        [62].13   // SPARE
        [60].8   // PANEL W3 SPONGE UNIT AUTO Sw. Pos.
        [60].9   // PANEL W3 SPONGE UNIT MANUAL Sw. Pos.
        [60].10   // PANEL W3 SPONGE UNIT ON Sw. Pos.
        [60].11   // PANEL W3 SPONGE UNIT OFF Sw. Pos.
        [60].12   // PANEL W3 AIR KNIFE AUTO Sw. Pos.
        [60].13   // PANEL W3 AIR KNIFE MANUAL Sw. Pos.
        [62].9   // SPARE
        [61].0   // PANEL W3 BRUSH #1 UPPER BRUSH CONVERGE Sw. Pos.
        [61].1   // PANEL W3 BRUSH #1 UPPER BRUSH RETRACT Sw. Pos.
        [61].4   // PANEL W3 SPONGE UNIT UPPER SPONGE CONVERGE Sw. Pos.
        [61].5   // PANEL W3 SPONGE UNIT UPPER SPONGE RETRACT Sw. Pos.
        [61].6   // PANEL W3 BRUSH #1 LOWER BRUSH CONVERGE Sw. Pos.
        [61].7   // PANEL W3 BRUSH #1 LOWER BRUSH RETRACT Sw. Pos.
        [61].10   // PANEL W3 SPONGE UNIT LOWER SPONGE CONVERGE Sw. Pos.
        [61].11   // PANEL W3 SPONGE UNIT LOWER SPONGE RETRACT Sw. Pos.
        [61].12   // PANEL W3 AIR KNIFE UNIT #1 CONVERGE Sw. Pos.
        [61].13   // PANEL W3 AIR KNIFE UNIT #1 RETRACT Sw. Pos.
        [61].14   // PANEL W3 AIR KNIFE UNIT #2 CONVERGE Sw. Pos.
        [61].15   // PANEL W3 AIR KNIFE UNIT #2 RETRACT Sw. Pos.
        [62].0   // PANEL W3 Cross break Reset Push-button
        [62].1   // PANEL W3 WATER SPRAYERS AUTO Sw. Pos.
        [62].2   // PANEL W3 WATER SPRAYERS MANUAL Sw. Pos.
        [62].3   // PANEL W3 WATER SPRAYERS ON Sw. Pos.
        [62].4   // PANEL W3 WATER SPRAYERS OFF Sw. Pos.
        [64].1   // VMCC M1 DC Input Power ON
        [64].2   // VMCC M1 DC Output Power ON
        [64].4   // VMCC M1 E-STOP Power ON
        [64].5   // VMCC M1 DC Power Supply #1 ON
        [64].6   // VMCC M1 DC Power Supply #2 ON
        [64].8   // VMCC M1 Alarm Silence
        [64].9   // VMCC M1 Alarm Reset
        [64].10   // VMCC M1 E-Stop Circuit Energized
        [64].11   // VMCC M1 Crusher Bar Lowered
        [64].12   // VMCC M1 Crusher Bar Raised
        [64].13   // VMCC M1 Crusher #1 Auto mode ON=AUTO OFF=MAN
        [64].14   // VMCC M1 Crusher #1 Manual raise
        [64].15   // VMCC M1 Crusher #1 Manual lower
        [65].0   // VMCC M1 Crusher #1 Drive Fault
        [65].1   // VMCC M1 Drive Alarm Light is ON
        [65].3   // VMCC M1 Crusher #1 Test Pushbutton
        [65].4   // No. 1 Crusher Chip Blower Start Pushbutton (Top)
        [65].5   // No. 1 Crusher Chip Blower Start Pushbutton (VMCC M1)
        [65].6   // No. 1 Crusher Chip Blower Stop Pushbutton (Top)
        [65].7   // No. 1 Crusher Chip Blower Stop Pushbutton (VMCC M1)
        [65].8   // VMCC M1 SPARE
        [65].12   // VMCC M1 Crusher #1 Start Pushbutton
        [65].13   // VMCC M1 Crusher #1 Stop Pushbutton
        [65].15   // VMCC M1 Generator Running bit
        [71].2   // MB -->> Cullet M47B Run Fwd Signal
        [71].3   // MB -->> Cullet M47B Run Rev Signal
        [80].0   // NO. 1 CRUSHER Signal from Reliance drive System E-STOP
        [80].1   // NO. 1 CRUSHER Signal from C.T. master drive System DRIVE FAULT
        [80].3   // IAL TEMPERATURE ALARM
        [80].4   // Lehr Conv AUX 1 Healthy Relay
        [80].5   // Lehr Conv AUX 2 Healthy Relay
        [80].6   // Lehr Conv AUX 3 Healthy Relay
        [80].7   // Lehr Conv AUX 4 Healthy Relay
        [80].8   // Lehr Conv AUX 5 Healthy Relay
        [80].9   // Lehr Conv AUX 6 Healthy Relay
        [80].10   // Lehr Conv AUX 7 Healthy Relay
        [80].11   // Lehr Conv AUX 8 Healthy Relay
        [80].12   // Lehr Conv AUX 9 Healthy Relay
        [80].13   // Lehr Conv AUX 10 Healthy Relay
        [80].14   // Lehr Conv AUX 11 Healthy Relay
        [80].15   // Lehr Conv AUX 12 Healthy Relay
        [81]   // AUTOMAX Lehr speed Received from AutoMax
        [83].0   // Lehr Conv AUX 13 Healthy Relay
        [83].1   // Lehr Conv AUX 14 Healthy Relay
        [83].2   // Lehr Conv AUX 15 Healthy Relay
        [83].3   // Lehr Conv AUX 16 Healthy Relay
        [83].4   // Lehr Conv AUX 17 Healthy Relay
        [112].1   // Cullet -->> MB M47B Conv Fwd Signal
        [112].2   // Cullet -->> MB M47B Conv Rev Signal
        [112].3   // Cullet -->> MB M37B Conv Fwd Signal
        [112].4   // Cullet -->> MB M37B Conv Rev Signal
        [113].1   // Cullet --> MB Panel C4 Equipment Fault or Failure
        [113].2   // Cullet --> MB Panel C1 Equipment Fault or Failure
        [113].3   // Cullet --> MB Panel C2 Equipment Fault or Failure
        [113].4   // Cullet --> MB Panel C3 Equipment Fault or Failure
        [121].1   // M2 -->> MB Crusher No. 4 Is Operating
        [121].2   // M2 -->> MB Crusher No. 3 is Operating
        [121].3   // M2 ---->> MB Crusher No. 2 Is Operating
        [123].0   // M2 -->> MB Drop #1 Crusher Pushbutton
        [123].1   // M2 -->> MB Trim deck E-stop
        [123].2   // M2 -->> MB Trim deck Drive system Critical Failure
        [123].3   // M2 -->> MB Trim deck Drive fault
        [123].4   // M2 -->> MB Mainline E-stop
        [123].6   // M2 -->> MB Mainline Drive fault
        [123].11   // M2 -->> MB Drive running M2CM01
        [123].12   // M2 -->> MB Mainline Backup to
        [123].13   // M2 -->> MB Crush-all Selector sw. Status
        [123].14   // M2 -->> MB Leg 2 Is In Sleep Mode Transfer Unavailable
        [123].15   // M2 -->> MB Leg 3 Is In Sleep Mode Transfer Unavailable
        [124].0   // M2 -->> MB Leg 4 Is In Sleep Mode Transfer Unavailable
        [124].1   // M2 -->> MB Leg 5 Is In Sleep Mode Transfer Unavailable
        [124].2   // M2 -->> MB ML is in Sleep Mode
        [124].3   // M2-->Mb UL Crusher Is Faulted
        [124].4   // M2-->MB VISION SYS Rejected Plate Alarm Horn
        [127].4   // M2-->MB Float Glass Prodution
        [123]   // M2 --> MB
        [65]   // VMCC M1 Crusher
        [113]   // Cullet --> MB
        [112]   // Cullet --> MB
        [64]   // VMCC M1 INPUTS
        [121].7   // M2 -->> MB ???
        [64].0   // VMCC M1 Drive Contactor Energized
        [28].13   // CRSSBRK ZONE 3 Adapter power ON
        [30].0   // CRSSBRK ZONE 4 North Outside Bypass Switch
        [28].14   // CRSSBRK ZONE 3 Input power ON
        [124]   // M2 --> MB
        [57]   // PANEL W2
        [34].10   // MANUAL INSPCTN MODE MAN
        [34].11   // MANUAL INSPCTN MODE AUTO
        [30].9   // IMAGE AUTO Retro Reflector
        [114]   // Cullet --> MB
        [115]   // Cullet --> MB
        [80]   // LEHR Conv Healthy Relays
        [116]   // Cullet --> MB
        [117]   // Cullet --> MB
        [56]   // PANEL W2
        [125]   // M2 --> MB
        [83]   // LEHR Conv Healthy Relays
        [118]   // Cullet --> MB
        [119]   // Cullet --> MB
        [43]   // VMCC W1
        [71]   // MB --> Cullet
        [42]   // VMCC W1
        [30]   // IMAGE AUTO CRSSBRK ZONE 4
        [32]   // APC CRSSBRK ZONE 5
        [18]   // APC
        [19]   // PROCESS STOP
        [121]   // M2 --> MB
        [61]   // PANEL W3
        [60]   // PANEL W3
        [30].6   // CRSSBRK ZONE 4 South Outside Photo-cell
        [30].7   // CRSSBRK ZONE 4 South Inside Photo-cell
        [30].8   // IMAGE AUTO Open Graticule Selector Switch (UP)
        [30].14   // IMAGE AUTO Close Graticule Selector Switch (DOWN)
        [30].11   // IMAGE AUTO Cover close Acknowledge Push-button (Silence)
        [34].2   // MANUAL INSPCTN Quality defect switch (Enable/Inhibit)
        [122]   // M2 --> MB
        [28]   // CRSSBRK ZONE 3
        [30].2   // CRSSBRK ZONE 4 South Outside Bypass Switch
        [30].3   // CRSSBRK ZONE 4 South Inside Bypass Switch
        [28].15   // CRSSBRK ZONE 3 Output power ON
        [30].4   // CRSSBRK ZONE 4 North Outside Photo-cell
        [56].14   // SPARE
        [127]   // M2 --> MB
        [26]   // CRSSBRK ZONE 2
        [126]   // M2 --> MB
        [17]   // Water
        [16]   // ISRA 5D
        [3]   // PROCESS STOP
        [24]   // CRSSBRK ZONE 1
        [62]   // PANEL W3
        [26].13   // CRSSBRK ZONE 2 Adapter power ON
        [33]   // APC
        [58]   // PANEL W2
        [12]   // Bridge
        [26].15   // CRSSBRK ZONE 2 Output power ON
        [26].14   // CRSSBRK ZONE 2 Input power ON
        [30].5   // CRSSBRK ZONE 4 North Inside Photo-cell
        [30].1   // CRSSBRK ZONE 4 North Inside Bypass Switch
        [18].0   // SPARE (MARKING BRIDGE On/Off Selector switch 0=off 1=on)
        [18].1   // SPARE (MARKING BRIDGE Auto/Manual 0=Manual 1=Auto)
        [16].2   // Spare
        [16].11   // Spare
        [16].12   // Spare
        [16].13   // Spare
        [16].15   // Spare
        [17].0   // Spare
        [17].6   // Spare
        [17].8   // Spare
        [17].12   // SPARE (Chilled Water Blower VFD Is At Speed)
        [17].15   // SPARE (ROCKWELL CAPPING SYSTEM: 50mm of Glass Travel Pulse Signal)
        [33].9   // SPARE (Apc system 0ff)
        [34]   // LOW-E MAUAL INSPCTN (MI_6CS)
        [43].4   // VMCC W1 Upper Sponge Drive fault (NOT USED ANYMORE)
        [43].5   // VMCC W1 Lower Sponge Drive fault (NOT USED ANYMORE)
        [42].1   // VMCC W1 Drive Contactor Energized (NOT USED ANYMORE)
        [42].2   // VMCC W1 DC Input Power ON (NOT USED ANYMORE)
        [42].3   // VMCC W1 DC Output Power ON (NOT USED ANYMORE)
        [42].5   // VMCC W1 E-STOP Power ON (NOT USED ANYMORE)
        [42].6   // VMCC W1 DC Power Supply #1 ON (NOT USED ANYMORE)
        [42].7   // VMCC W1 DC Power Supply #2 ON (NOT USED ANYMORE)
        [42].8   // VMCC W1 Alarm Silence (NOT USED ANYMORE)
        [42].10   // VMCC W1 E-STOP ACTIVE (NOT USED ANYMORE)
        [42].11   // VMCC W1 Drive Comm. Power (NOT USED ANYMORE)
        [43].12   // VMCC W1 Crusher #1 Start Pushbutton (NOT USED ANYMORE)
        [43].13   // VMCC W1 Crusher #1 Stop Pushbutton (NOT USED ANYMORE)
        [56].4   // PANEL W2 BRUSH #2 AUTO Sw. Pos. (NOT USED ANYMORE)
        [56].5   // PANEL W2 BRUSH #2 MANUAL Sw. Pos. (NOT USED ANYMORE)
        [56].6   // PANEL W2 BRUSH #2 ON Sw. Pos. (NOT USED ANYMORE)
        [56].7   // PANEL W2 BRUSH #2 OFF Sw. Pos. (NOT USED ANYMORE)
        [57].2   // PANEL W2 BRUSH #2 UPPER BRUSH CONVERGE Sw. Pos. (NOT USED ANYMORE)
        [57].3   // PANEL W2 BRUSH #2 UPPER BRUSH RETRACT Sw. Pos. (NOT USED ANYMORE)
        [57].8   // PANEL W2 BRUSH #2 LOWER BRUSH CONVERGE Sw. Pos. (NOT USED ANYMORE)
        [57].9   // PANEL W2 BRUSH #2 LOWER BRUSH RETRACT Sw. Pos. (NOT USED ANYMORE)
        [60].4   // PANEL W3 BRUSH #2 AUTO Sw. Pos. (NOT USED ANYMORE)
        [60].5   // PANEL W3 BRUSH #2 MANUAL Sw. Pos. (NOT USED ANYMORE)
        [60].6   // PANEL W3 BRUSH #2 ON Sw. Pos. (NOT USED ANYMORE)
        [60].7   // PANEL W3 BRUSH #2 OFF Sw. Pos. (NOT USED ANYMORE)
        [61].2   // PANEL W3 BRUSH #2 UPPER BRUSH CONVERGE Sw. Pos. (NOT USED ANYMORE)
        [61].3   // PANEL W3 BRUSH #2 UPPER BRUSH RETRACT Sw. Pos. (NOT USED ANYMORE)
        [61].8   // PANEL W3 BRUSH #2 LOWER BRUSH CONVERGE Sw. Pos. (NOT USED ANYMORE)
        [61].9   // PANEL W3 BRUSH #2 LOWER BRUSH RETRACT Sw. Pos. (NOT USED ANYMORE)
        [58].5   // PANEL W2 SELECTOR SWITCH CITRIC ACID WASHER ON (# W2) (NOT USED ANYMORE)
        [58].6   // PANEL W2 SELECTOR SWITCH CITRIC ACID WASHER OFF (# W2) (NOT USED ANYMORE)
        [62].5   // PANEL W3 SELECTOR SWITCH CITRIC ACID WASHER ON (# W3) (NOT USED ANYMORE)
        [62].6   // PANEL W3 SELECTOR SWITCH CITRIC ACID WASHER OFF (# W3) (NOT USED ANYMORE)
        [113].0   // Cullet --> MB SYSTEM LOCAL HEARTBEAT FOR HOST PLC
        [113].5   // Cullet --> MB FIX MMI M-47B Conveyor Running Reverse
        [114].1   // LEG 4 EOL FEEDER AUTO RUN STATUS
        [114].2   // LEG 5 EOL FEEDER AUTO RUN STATUS
        [114].3   // PANEL C4 - TRIM DROP VP 917078 Running at Speed
        [114].4   // PANEL C3 - CR#3 VP 917067 VFD FAULT STATUS
        [114].5   // PANEL C3 - CR#3 VP 917067 VFD RUNNING STATUS
        [114].6   // PANEL C3 M34T TO M34 TRANS VP 917066 VFD FAULT STATUS
        [114].7   // PANEL C3 M34T TO M34 TRANS VP 917066 VFD RUNNING STATUS
        [114].10   // PANEL C3 VP 917070 VFD FAULT STATUS
        [114].11   // PANEL C3 VP 917070 VFD RUNNING STATUS
        [114].12   // PANEL C3 VP 917071 VFD FAULT STATUS
        [114].13   // PANEL C3 VP 917071 VFD RUNNING STATUS
        [114].14   // PANEL C2 VP 917077 VFD FAULT STATUS
        [114].15   // PANEL C2 VP 917077 VFD RUNNING STATUS
        [115].0   // PANEL C4 M34T MAIN #1 CONV RUNNING STATUS
        [115].1   // LEG 3 EOL FEEDER AUTO RUN STATUS
        [115].2   // PANEL C4 M-32 CONVEYOR RUNNING STATUS
        [115].3   // PANEL C4 M-33 CONVEYOR RUNNING STATUS
        [115].4   // PANEL C4 M34T MAIN #1 CONV E-STOP STATUS
        [115].6   // PANEL C4 M-32 CONVEYOR E-STOP STATUS
        [115].7   // PANEL C4 M-33 CONVEYOR E-STOP STATUS
        [115].8   // PANEL C4 M34T MAIN CONV #1 ZERO SPEED STATUS
        [115].10   // PANEL C4 M-32 CONVEYOR ZERO SPEED SWITCH STATUS
        [115].11   // PANEL C4 M-33 CONVEYOR ZERO SPEED STATUS
        [115].12   // PANEL C2 VP 917076 VFD FAULT STATUS
        [115].13   // PANEL C2 VP 917076 VFD RUNNING STATUS
        [115].14   // PANEL C2 VP 917075 VFD FAULT STATUS
        [115].15   // PANEL C2 VP 917075 VFD RUNNING STATUS
        [116].0   // PANEL C4 - CR#4 VP 917068 VFD RUNNING STATUS
        [116].1   // LEG 5 FEEDER DRIVE RUNNING STATUS
        [116].2   // PANEL C2 VP 917074 VFD FAULT STATUS
        [116].3   // PANEL C2 VP 917074 VFD RUNNING STATUS
        [116].4   // PANEL C4 - CR#4 VP 917068 VFD FAULT STATUS
        [116].7   // PANEL C2 VP 917073 VFD FAULT STATUS
        [116].8   // PANEL C2 VP 917073 VFD RUNNING STATUS
        [116].9   // PANEL C2 VP 917072 VFD FAULT STATUS
        [116].10   // PANEL C2 VP 917072 VFD RUNNING STATUS
        [116].11   // PANEL C1 VP 917060 VFD FAULT STATUS
        [116].12   // PANEL C1 VP 917060 VFD RUNNING STATUS
        [116].13   // PANEL C3 M-40 CONVEYOR RUNNING STATUS
        [116].14   // PANEL C3 M-40 CONVEYOR E-STOP STATUS
        [116].15   // PANEL C3 M-40 CONVEYOR ZERO SPEED SWITCH STATUS
        [117].0   // M47A_RUN_STAT PANEL C1 M-47A CONVEYOR RUNNING STATUS
        [117].1   // M47A_ESTOP_STAT PANEL C1 M-47A CONVEYOR E-STOP STATUS
        [117].2   // M47A_ZSS_STAT PANEL C1 M-47A CONVEYOR ZERO SPEED SWITCH STATUS
        [117].3   // M47B_RUN_STAT PANEL C1 M-47B CONVEYOR RUNNING STATUS
        [117].4   // M47B_ESTOP_STAT PANEL C1 M-47B CONVEYOR E-STOP STATUS
        [117].5   // M47B_ZSS_STAT PANEL C1 M-47B CONVEYOR ZERO SPEED SWITCH STATUS
        [117].6   // M46_RUN_STAT PANEL C1 M-46 CONVEYOR RUNNING STATUS
        [117].7   // M46_ESTOP_STAT PANEL C1 M-46 CONVEYOR E-STOP STATUS
        [117].8   // M46_ZSS_STAT PANEL C1 M-46 CONVEYOR ZERO SPEED SWITCH STATUS
        [117].9   // M45B_RUN_STAT PANEL C1 M-45B CONVEYOR RUNNING STATUS
        [117].10   // M45B_ESTOP_STAT PANEL C1 M-45B CONVEYOR E-STOP STATUS
        [117].11   // M45B_ZSS_STAT PANEL C1 M-45B CONVEYOR ZERO SPEED SWITCH STATUS
        [117].12   // M37A_RUN_STAT PANEL C2 M-37A CONVEYOR RUNNING STATUS
        [117].13   // M37A_ESTOP_STAT PANEL C2 M-37A CONVEYOR E-STOP STATUS
        [117].14   // M37A_ZSS_STAT PANEL C2 M-37A CONVEYOR ZERO SPEED SWITCH STATUS
        [117].15   // M37B_RUN_STAT PANEL C2 M-37B CONVEYOR RUNNING STATUS
        [118].0   // M37B_ESTOP_STAT PANEL C2 M-37B CONVEYOR E-STOP STATUS
        [118].1   // M37B_ZSS_STAT PANEL C2 M-37B CONVEYOR ZERO SPEED SWITCH STATUS
        [118].2   // M36_RUN_STAT PANEL C2 M-36 CONVEYOR RUNNING STATUS
        [118].3   // M36_ESTOP_STAT PANEL C2 M-36 CONVEYOR E-STOP STATUS
        [118].4   // M36_ZSS_STAT PANEL C2 M-36 CONVEYOR ZERO SPEED SWITCH STATUS
        [118].5   // M35_RUN_STAT PANEL C2 M-35 CONVEYOR RUNNING STATUS
        [118].6   // M35_ESTOP_STAT PANEL C2 M-35 CONVEYOR E-STOP STATUS
        [118].7   // M35_ZSS_STAT PANEL C2 M-35 CONVEYOR ZERO SPEED SWITCH STATUS
        [118].8   // CHPR_RUN_STAT PANEL C2 CHOPPER 917014 RUNNING STATUS
        [118].9   // CHPR_ESTOP_STAT PANEL C2 CHOPPER 917014 E-STOP STATUS
        [118].10   // CHPR_ZSS_STAT PANEL C2 CHOPPER 917014 ZERO SPEED SWITCH STATUS
        [118].11   // M45_RUN_STAT PANEL C2 M-45 CONVEYOR RUNNING STATUS
        [118].12   // M45_ESTOP_STAT PANEL C2 M-45 CONVEYOR E-STOP STATUS
        [118].13   // M45_ZSS_STAT PANEL C2 M-45 CONVEYOR ZERO SPEED SWITCH STATUS
        [118].14   // M45A_RUN_STAT PANEL C2 M-45A CONVEYOR RUNNING STATUS
        [118].15   // M45A_ESTOP_STAT PANEL C2 M-45A CONVEYOR E-STOP STATUS
        [119].0   // M45A_ZSS_STAT PANEL C2 M-45A CONVEYOR ZERO SPEED SWITCH STATUS
        [119].1   // M34_RUN_STAT PANEL C3 M-34 CONVEYOR RUNNING STATUS
        [119].2   // M34_ESTOP_STAT PANEL C3 M-34 CONVEYOR E-STOP STATUS
        [119].3   // M34_ZSS_STAT PANEL C3 M-34 CONVEYOR ZERO SPEED SWITCH STATUS
        [119].4   // M44_RUN_STAT PANEL C3 M-44 CONVEYOR RUNNING STATUS
        [119].5   // M44_ESTOP_STAT PANEL C3 M-44 CONVEYOR E-STOP STATUS
        [119].6   // M44_ZSS_STAT PANEL C3 M-44 CONVEYOR ZERO SPEED SWITCH STATUS
        [119].7   // M43_RUN_STAT PANEL C3 M-43 CONVEYOR RUNNING STATUS
        [119].8   // M43_ESTOP_STAT PANEL C3 M-43 CONVEYOR E-STOP STATUS
        [119].9   // M43_ZSS_STAT PANEL C3 M-43 CONVEYOR ZERO SPEED SWITCH STATUS
        [119].10   // M41_RUN_STAT PANEL C3 M-41 CONVEYOR RUNNING STATUS
        [119].11   // M41_ESTOP_STAT PANEL C3 M-41 CONVEYOR E-STOP STATUS
        [119].12   // M41_ZSS_STAT PANEL C3 M-41 CONVEYOR ZERO SPEED SWITCH STATUS
        [119].13   // M42_RUN_STAT PANEL C3 M-42 CONVEYOR RUNNING STATUS
        [119].14   // M42_ESTOP_STAT PANEL C3 M-42 CONVEYOR E-STOP STATUS
        [119].15   // M42_ZSS_STAT PANEL C3 M-42 CONVEYOR ZERO SPEED SWITCH STATUS
   IA_ACK_PB : ALIAS FOR I[30].11;
   IA_CLOSE_GRAT : ALIAS FOR I[30].14;
   IA_COVER_CLOSED : ALIAS FOR N54[281].5;
   IA_COVER_VLVE : ALIAS FOR O[31].10;
   IA_GRAT_OPEN_SS : ALIAS FOR I[30].8;
   IA_RET_CL_PROX : ALIAS FOR I[30].12;
   IA_RET_CLSD_ACK : ALIAS FOR N54[281].6;
   INDEX : ALIAS FOR S[24];
   INIT_TIMER : ALIAS FOR T4[0];
   IW_FE1_BTR : ALIAS FOR W_N7[32];
   LEG2_SLEEP : ALIAS FOR I[123].14;
   LEG3_SLEEP : ALIAS FOR I[123].15;
   LEG4_SLEEP : ALIAS FOR I[124].0;
   LEG5_SLEEP : ALIAS FOR I[124].1;
   LEHR_2IN_PULSE : ALIAS FOR B73[0].1;
   LEHR_SPEED : ALIAS FOR N60[1];
   LEHRSPD_AUTOMAX : ALIAS FOR N98[1];
   LEHRSPD_AVE : ALIAS FOR N98[2];
   LEHRSPD_CURRENT : ALIAS FOR N98[5];
   LEHRSPD_STD : ALIAS FOR N98[3];
   M1_ALM_FLT_RLY : ALIAS FOR O[66].13;
   M1_ALM_RESET : ALIAS FOR I[64].9;
   M1_ALM_SILENCE : ALIAS FOR I[64].8;
   M1_DC_INPOW : ALIAS FOR I[64].1;
   M1_DC_OUTPOW : ALIAS FOR I[64].2;
   M1_DC_PS1 : ALIAS FOR I[64].5;
   M1_DC_PS2 : ALIAS FOR I[64].6;
   M1_DRV_CONT_ON : ALIAS FOR I[64].0;
   M1_ESTOP_ON : ALIAS FOR I[64].10;
   M1_ESTOPPOW : ALIAS FOR I[64].4;
   M202_M1_DR : AXIS_CIP_DRIVE; {access Read Only}
   M202_M1_DR_IN_MAJ : MOTION_INSTRUCTION := (FLAGS := 570425344, DN := 1); {access None}
   M202_M1_DR_IN_MAM : MOTION_INSTRUCTION := (FLAGS := 33554432); {access None}
   M202_M1_DR_IN_MAR : MOTION_INSTRUCTION := (FLAGS := 33554432); {access None}
   M202_M1_DR_IN_MAS : MOTION_INSTRUCTION := (FLAGS := -1442840576, EN := 1, DN := 1, PC := 1); {access None}
   M202_M1_DR_IN_MCD : MOTION_INSTRUCTION := (FLAGS := 570425344, DN := 1); {access None}
   M202_M1_DR_IN_MRP : MOTION_INSTRUCTION := (FLAGS := 33554432); {access None}
   M202_M1_DR_MAFR : MOTION_INSTRUCTION := (FLAGS := 301989888, ER := 1, ERR := 11); {access None}
   M202_M1_DR_MDR : MOTION_INSTRUCTION := (FLAGS := -1845493760, EN := 1, ER := 1, ERR := 11); {access None}
   M202_M1_DR_MSF : MOTION_INSTRUCTION := (FLAGS := 570425344, DN := 1, STATUS := 2, STATE := 1); {access None}
   M202_M1_DR_MSO : MOTION_INSTRUCTION := (FLAGS := -1610612736, EN := 1, DN := 1, STATE := 1); {access None}
   M202_M1_DR_OUT_MAJ : MOTION_INSTRUCTION := (FLAGS := 570425344, DN := 1); {access None}
   M202_M1_DR_OUT_MAM : MOTION_INSTRUCTION := (FLAGS := 33554432); {access None}
   M202_M1_DR_OUT_MAR : MOTION_INSTRUCTION := (FLAGS := 33554432); {access None}
   M202_M1_DR_OUT_MAS : MOTION_INSTRUCTION := (FLAGS := -1442840576, EN := 1, DN := 1, PC := 1); {access None}
   M202_M1_DR_OUT_MCD : MOTION_INSTRUCTION := (FLAGS := 570425344, DN := 1); {access None}
   M202_M1_DR_OUT_MRP : MOTION_INSTRUCTION := (FLAGS := 33554432); {access None}
   M203_M1_DR : AXIS_CIP_DRIVE; {access Read Only}
   M203_M1_DR_IN_MAJ : MOTION_INSTRUCTION := (FLAGS := 570425344, DN := 1); {access None}
   M203_M1_DR_IN_MAM : MOTION_INSTRUCTION := (FLAGS := 33554432); {access None}
   M203_M1_DR_IN_MAR : MOTION_INSTRUCTION := (FLAGS := 33554432); {access None}
   M203_M1_DR_IN_MAS : MOTION_INSTRUCTION := (FLAGS := -1442840576, EN := 1, DN := 1, PC := 1); {access None}
   M203_M1_DR_IN_MCD : MOTION_INSTRUCTION := (FLAGS := 570425344, DN := 1); {access None}
   M203_M1_DR_IN_MRP : MOTION_INSTRUCTION := (FLAGS := 33554432); {access None}
   M203_M1_DR_MAFR : MOTION_INSTRUCTION := (FLAGS := 301989888, ER := 1, ERR := 11); {access None}
   M203_M1_DR_MDR : MOTION_INSTRUCTION := (FLAGS := -1845493760, EN := 1, ER := 1, ERR := 11); {access None}
   M203_M1_DR_MSF : MOTION_INSTRUCTION := (FLAGS := 570425344, DN := 1, STATUS := 2, STATE := 1); {access None}
   M203_M1_DR_MSO : MOTION_INSTRUCTION := (FLAGS := -1610612736, EN := 1, DN := 1, STATE := 1); {access None}
   M203_M1_DR_OUT_MAJ : MOTION_INSTRUCTION := (FLAGS := 570425344, DN := 1); {access None}
   M203_M1_DR_OUT_MAM : MOTION_INSTRUCTION := (FLAGS := 33554432); {access None}
   M203_M1_DR_OUT_MAR : MOTION_INSTRUCTION := (FLAGS := 33554432); {access None}
   M203_M1_DR_OUT_MAS : MOTION_INSTRUCTION := (FLAGS := -1442840576, EN := 1, DN := 1, PC := 1); {access None}
   M203_M1_DR_OUT_MCD : MOTION_INSTRUCTION := (FLAGS := 570425344, DN := 1); {access None}
   M203_M1_DR_OUT_MRP : MOTION_INSTRUCTION := (FLAGS := 33554432); {access None}
   M203DROP : MAC_DROPCONV := (OUTPUT_xHLUpDownPushbutton := 1, INPUT_xProtection := 1, INPUT_xProtectionBrake := 1, AUX_tmOFFEachCutAcceleration.PRE := 2000, AUX_tmOFFEachCutAcceleration.ACC := 2000, AUX_tmOFFAcceleration.PRE := 8805, AUX_tmOFFAcceleration.ACC := 8805, AUX_tmONFeedbackMovAlarm.PRE := 2000, AUX_tmONFeedbackAlarm.PRE := 2000, AUX_tmONFeedbackBrakeAlarm.PRE := 7000, AUX_tmONMismatchSensorAlarm.PRE := 7000, AUX_tmONUpSensorAlarm.PRE := 5000, AUX_tmONDownSensorAlarm.PRE := 5000, AUX_tmONForceUp.PRE := 2000, AUX_tmONEmCutTimeout.PRE := 120000, AUX_dDistanceToDescent_cmm := 25000, AUX_dDistanceToCheckGlass_cmm := 100000, AUX_dConveyorLength_cmm := 440000, AUX_dAccelerationTime_ms := 2147483647, AUX_dAccelerationFactor := 3, AUX_dMaxSpeed_mm_min := 30000, ST_xConveyorDwRequest := 1, OSR_xCutForQltPopupEnd := 1); {access None}
   M203DROP_ALM : MAC_DROPCONV_ALM; {access Read Only}
        .rgxStoppingFaults[0].0   // Protection lifting
        .rgxStoppingFaults[0].1   // Protection brake
        .rgxStoppingFaults[0].2   // Feedback lifting
        .rgxStoppingFaults[0].3   // Feedback brake
        .rgxStoppingFaults[0].5   // A206SQ2.Timeout frame low
        .rgxStoppingFaults[0].6   // A206SQ1/2.Sensor high/low mismatch (same status)
        .rgxStoppingFaults[0].4   // A206SQ1.Timeout frame high
        .rgxStoppingFaults[0].7   // A206SQ3/4.Tilting safety bar disinsered
   M203DROP_HMR : MAC_DROPCONV_HMR := (dMode := 1, dStatus := 1, dDistanceFromSnaproll_cmm := 4190000); {access Read Only}
   M203DROP_HMW : MAC_DROPCONV_HMW := (dDistanceFromSnaproll_cmm := 4632000);
   M204_M1_DR : AXIS_CIP_DRIVE; {access Read Only}
   M204_M1_DR_IN_MAJ : MOTION_INSTRUCTION := (FLAGS := 570425344, DN := 1); {access None}
   M204_M1_DR_IN_MAM : MOTION_INSTRUCTION := (FLAGS := 33554432); {access None}
   M204_M1_DR_IN_MAR : MOTION_INSTRUCTION := (FLAGS := 33554432); {access None}
   M204_M1_DR_IN_MAS : MOTION_INSTRUCTION := (FLAGS := -1442840576, EN := 1, DN := 1, PC := 1); {access None}
   M204_M1_DR_IN_MCD : MOTION_INSTRUCTION := (FLAGS := 570425344, DN := 1); {access None}
   M204_M1_DR_IN_MRP : MOTION_INSTRUCTION := (FLAGS := 33554432); {access None}
   M204_M1_DR_MAFR : MOTION_INSTRUCTION := (FLAGS := 301989888, ER := 1, ERR := 11); {access None}
   M204_M1_DR_MDR : MOTION_INSTRUCTION := (FLAGS := -1845493760, EN := 1, ER := 1, ERR := 11); {access None}
   M204_M1_DR_MSF : MOTION_INSTRUCTION := (FLAGS := 570425344, DN := 1, STATUS := 2, STATE := 1); {access None}
   M204_M1_DR_MSO : MOTION_INSTRUCTION := (FLAGS := -1610612736, EN := 1, DN := 1, STATE := 1); {access None}
   M204_M1_DR_OUT_MAJ : MOTION_INSTRUCTION := (FLAGS := 570425344, DN := 1); {access None}
   M204_M1_DR_OUT_MAM : MOTION_INSTRUCTION := (FLAGS := 33554432); {access None}
   M204_M1_DR_OUT_MAR : MOTION_INSTRUCTION := (FLAGS := 33554432); {access None}
   M204_M1_DR_OUT_MAS : MOTION_INSTRUCTION := (FLAGS := -1442840576, EN := 1, DN := 1, PC := 1); {access None}
   M204_M1_DR_OUT_MCD : MOTION_INSTRUCTION := (FLAGS := 570425344, DN := 1); {access None}
   M204_M1_DR_OUT_MRP : MOTION_INSTRUCTION := (FLAGS := 33554432); {access None}
   M205BREAKER : MAC_BREAKER := (ST_xBreakerRunningRequest := 1, OSR_xBreakerRunning := 1, INPUT_xProtectionFan := 1, INPUT_xStopBreaker := 1, INPUT_xThermalProbe := 1, OUTPUT_xBreakerRun := 1, AUX_tmONCrusherStopDelayed.PRE := 320000, AUX_tmONFeedbackBreakerRot.PRE := 15000, AUX_tmONBreakControlRotation.PRE := 5000, AUX_tmONFeedbackBrakeBreakRot.PRE := 2000, AUX_tmONFeedbackExclusionInduct.PRE := 5000); {access None}
   M205BREAKER_ALM : MAC_BREAKER_ALM; {access Read Only}
        .rgxStoppingFaults[0].5   // Exclusion inductance feedback
        .rgxStoppingFaults[0].3   // Drive error
        .rgdCodeAlarm[0]   // A60AZ1.Error Code
        .rgxStoppingFaults[0].2   // Motor thermal probe
        .rgxStoppingFaults[0].4   // A56QS1.Safety motor sectioning
        .rgxStoppingFaults[0].0   // Rotation feedback
        .rgxStoppingFaults[0].1   // Protection rotation
        .rgxStoppingFaults[0].6   // A207SQ1.Breaker rotation sensor
        .rgxFaults[0].0   // A63QM2.Protection fan rotation
   M205BREAKER_HMR : MAC_BREAKER_HMR := (dBreakerStatus := 1); {access Read Only}
   M205BREAKER_HMW : MAC_BREAKER_HMW := (dTimeoutRunningCrusher_ms := 320000);
   M206_M1_DR : AXIS_CIP_DRIVE; {access Read Only}
   M206_M1_DR_IN_MAJ : MOTION_INSTRUCTION := (FLAGS := 570425344, DN := 1); {access None}
   M206_M1_DR_IN_MAM : MOTION_INSTRUCTION := (FLAGS := 33554432); {access None}
   M206_M1_DR_IN_MAR : MOTION_INSTRUCTION := (FLAGS := 33554432); {access None}
   M206_M1_DR_IN_MAS : MOTION_INSTRUCTION := (FLAGS := -1442840576, EN := 1, DN := 1, PC := 1); {access None}
   M206_M1_DR_IN_MCD : MOTION_INSTRUCTION := (FLAGS := 570425344, DN := 1); {access None}
   M206_M1_DR_IN_MRP : MOTION_INSTRUCTION := (FLAGS := 33554432); {access None}
   M206_M1_DR_MAFR : MOTION_INSTRUCTION := (FLAGS := 301989888, ER := 1, ERR := 11); {access None}
   M206_M1_DR_MDR : MOTION_INSTRUCTION := (FLAGS := -1845493760, EN := 1, ER := 1, ERR := 11); {access None}
   M206_M1_DR_MSF : MOTION_INSTRUCTION := (FLAGS := 570425344, DN := 1, STATUS := 2, STATE := 1); {access None}
   M206_M1_DR_MSO : MOTION_INSTRUCTION := (FLAGS := -1610612736, EN := 1, DN := 1, STATE := 1); {access None}
   M206_M1_DR_OUT_MAJ : MOTION_INSTRUCTION := (FLAGS := 570425344, DN := 1); {access None}
   M206_M1_DR_OUT_MAM : MOTION_INSTRUCTION := (FLAGS := 33554432); {access None}
   M206_M1_DR_OUT_MAR : MOTION_INSTRUCTION := (FLAGS := 33554432); {access None}
   M206_M1_DR_OUT_MAS : MOTION_INSTRUCTION := (FLAGS := -1442840576, EN := 1, DN := 1, PC := 1); {access None}
   M206_M1_DR_OUT_MCD : MOTION_INSTRUCTION := (FLAGS := 570425344, DN := 1); {access None}
   M206_M1_DR_OUT_MRP : MOTION_INSTRUCTION := (FLAGS := 33554432); {access None}
   M207_M1_DR : AXIS_CIP_DRIVE; {access Read Only}
   M207_M1_DR_IN_MAJ : MOTION_INSTRUCTION := (FLAGS := 570425344, DN := 1); {access None}
   M207_M1_DR_IN_MAM : MOTION_INSTRUCTION := (FLAGS := 33554432); {access None}
   M207_M1_DR_IN_MAR : MOTION_INSTRUCTION := (FLAGS := 33554432); {access None}
   M207_M1_DR_IN_MAS : MOTION_INSTRUCTION := (FLAGS := -1442840576, EN := 1, DN := 1, PC := 1); {access None}
   M207_M1_DR_IN_MCD : MOTION_INSTRUCTION := (FLAGS := 570425344, DN := 1); {access None}
   M207_M1_DR_IN_MRP : MOTION_INSTRUCTION := (FLAGS := 33554432); {access None}
   M207_M1_DR_MAFR : MOTION_INSTRUCTION := (FLAGS := 301989888, ER := 1, ERR := 11); {access None}
   M207_M1_DR_MDR : MOTION_INSTRUCTION := (FLAGS := -1845493760, EN := 1, ER := 1, ERR := 11); {access None}
   M207_M1_DR_MSF : MOTION_INSTRUCTION := (FLAGS := 570425344, DN := 1, STATUS := 2, STATE := 1); {access None}
   M207_M1_DR_MSO : MOTION_INSTRUCTION := (FLAGS := -1610612736, EN := 1, DN := 1, STATE := 1); {access None}
   M207_M1_DR_OUT_MAJ : MOTION_INSTRUCTION := (FLAGS := 570425344, DN := 1); {access None}
   M207_M1_DR_OUT_MAM : MOTION_INSTRUCTION := (FLAGS := 33554432); {access None}
   M207_M1_DR_OUT_MAR : MOTION_INSTRUCTION := (FLAGS := 33554432); {access None}
   M207_M1_DR_OUT_MAS : MOTION_INSTRUCTION := (FLAGS := -1442840576, EN := 1, DN := 1, PC := 1); {access None}
   M207_M1_DR_OUT_MCD : MOTION_INSTRUCTION := (FLAGS := 570425344, DN := 1); {access None}
   M207_M1_DR_OUT_MRP : MOTION_INSTRUCTION := (FLAGS := 33554432); {access None}
   M208_M1_DR : AXIS_CIP_DRIVE; {access Read Only}
   M208_M1_DR_IN_MAJ : MOTION_INSTRUCTION := (FLAGS := 570425344, DN := 1); {access None}
   M208_M1_DR_IN_MAM : MOTION_INSTRUCTION := (FLAGS := 33554432); {access None}
   M208_M1_DR_IN_MAR : MOTION_INSTRUCTION := (FLAGS := 33554432); {access None}
   M208_M1_DR_IN_MAS : MOTION_INSTRUCTION := (FLAGS := -1442840576, EN := 1, DN := 1, PC := 1); {access None}
   M208_M1_DR_IN_MCD : MOTION_INSTRUCTION := (FLAGS := 570425344, DN := 1); {access None}
   M208_M1_DR_IN_MRP : MOTION_INSTRUCTION := (FLAGS := 33554432); {access None}
   M208_M1_DR_MAFR : MOTION_INSTRUCTION := (FLAGS := 301989888, ER := 1, ERR := 11); {access None}
   M208_M1_DR_MDR : MOTION_INSTRUCTION := (FLAGS := -1845493760, EN := 1, ER := 1, ERR := 11); {access None}
   M208_M1_DR_MSF : MOTION_INSTRUCTION := (FLAGS := 570425344, DN := 1, STATUS := 2, STATE := 1); {access None}
   M208_M1_DR_MSO : MOTION_INSTRUCTION := (FLAGS := -1610612736, EN := 1, DN := 1, STATE := 1); {access None}
   M208_M1_DR_OUT_MAJ : MOTION_INSTRUCTION := (FLAGS := 570425344, DN := 1); {access None}
   M208_M1_DR_OUT_MAM : MOTION_INSTRUCTION := (FLAGS := 33554432); {access None}
   M208_M1_DR_OUT_MAR : MOTION_INSTRUCTION := (FLAGS := 33554432); {access None}
   M208_M1_DR_OUT_MAS : MOTION_INSTRUCTION := (FLAGS := -1442840576, EN := 1, DN := 1, PC := 1); {access None}
   M208_M1_DR_OUT_MCD : MOTION_INSTRUCTION := (FLAGS := 570425344, DN := 1); {access None}
   M208_M1_DR_OUT_MRP : MOTION_INSTRUCTION := (FLAGS := 33554432); {access None}
   M209_M1_DR : AXIS_CIP_DRIVE; {access Read Only}
   M209_M1_DR_IN_MAJ : MOTION_INSTRUCTION := (FLAGS := 570425344, DN := 1); {access None}
   M209_M1_DR_IN_MAM : MOTION_INSTRUCTION := (FLAGS := 33554432); {access None}
   M209_M1_DR_IN_MAR : MOTION_INSTRUCTION := (FLAGS := 33554432); {access None}
   M209_M1_DR_IN_MAS : MOTION_INSTRUCTION := (FLAGS := -1442840576, EN := 1, DN := 1, PC := 1); {access None}
   M209_M1_DR_IN_MCD : MOTION_INSTRUCTION := (FLAGS := 570425344, DN := 1); {access None}
   M209_M1_DR_IN_MRP : MOTION_INSTRUCTION := (FLAGS := 33554432); {access None}
   M209_M1_DR_MAFR : MOTION_INSTRUCTION := (FLAGS := 301989888, ER := 1, ERR := 11); {access None}
   M209_M1_DR_MDR : MOTION_INSTRUCTION := (FLAGS := -1845493760, EN := 1, ER := 1, ERR := 11); {access None}
   M209_M1_DR_MSF : MOTION_INSTRUCTION := (FLAGS := 570425344, DN := 1, STATUS := 2, STATE := 1); {access None}
   M209_M1_DR_MSO : MOTION_INSTRUCTION := (FLAGS := -1610612736, EN := 1, DN := 1, STATE := 1); {access None}
   M209_M1_DR_OUT_MAJ : MOTION_INSTRUCTION := (FLAGS := 570425344, DN := 1); {access None}
   M209_M1_DR_OUT_MAM : MOTION_INSTRUCTION := (FLAGS := 33554432); {access None}
   M209_M1_DR_OUT_MAR : MOTION_INSTRUCTION := (FLAGS := 33554432); {access None}
   M209_M1_DR_OUT_MAS : MOTION_INSTRUCTION := (FLAGS := -1442840576, EN := 1, DN := 1, PC := 1); {access None}
   M209_M1_DR_OUT_MCD : MOTION_INSTRUCTION := (FLAGS := 570425344, DN := 1); {access None}
   M209_M1_DR_OUT_MRP : MOTION_INSTRUCTION := (FLAGS := 33554432); {access None}
   M210_M1_DR : AXIS_CIP_DRIVE; {access Read Only}
   M210_M1_DR_IN_MAJ : MOTION_INSTRUCTION := (FLAGS := 570425344, DN := 1); {access None}
   M210_M1_DR_IN_MAM : MOTION_INSTRUCTION := (FLAGS := 33554432); {access None}
   M210_M1_DR_IN_MAR : MOTION_INSTRUCTION := (FLAGS := 33554432); {access None}
   M210_M1_DR_IN_MAS : MOTION_INSTRUCTION := (FLAGS := -1442840576, EN := 1, DN := 1, PC := 1); {access None}
   M210_M1_DR_IN_MCD : MOTION_INSTRUCTION := (FLAGS := 570425344, DN := 1); {access None}
   M210_M1_DR_IN_MRP : MOTION_INSTRUCTION := (FLAGS := 33554432); {access None}
   M210_M1_DR_MAFR : MOTION_INSTRUCTION := (FLAGS := 301989888, ER := 1, ERR := 11); {access None}
   M210_M1_DR_MDR : MOTION_INSTRUCTION := (FLAGS := -1845493760, EN := 1, ER := 1, ERR := 11); {access None}
   M210_M1_DR_MSF : MOTION_INSTRUCTION := (FLAGS := 570425344, DN := 1, STATUS := 2, STATE := 1); {access None}
   M210_M1_DR_MSO : MOTION_INSTRUCTION := (FLAGS := -1610612736, EN := 1, DN := 1, STATE := 1); {access None}
   M210_M1_DR_OUT_MAJ : MOTION_INSTRUCTION := (FLAGS := 570425344, DN := 1); {access None}
   M210_M1_DR_OUT_MAM : MOTION_INSTRUCTION := (FLAGS := 33554432); {access None}
   M210_M1_DR_OUT_MAR : MOTION_INSTRUCTION := (FLAGS := 33554432); {access None}
   M210_M1_DR_OUT_MAS : MOTION_INSTRUCTION := (FLAGS := -1442840576, EN := 1, DN := 1, PC := 1); {access None}
   M210_M1_DR_OUT_MCD : MOTION_INSTRUCTION := (FLAGS := 570425344, DN := 1); {access None}
   M210_M1_DR_OUT_MRP : MOTION_INSTRUCTION := (FLAGS := 33554432); {access None}
   M211_M1_DR : AXIS_CIP_DRIVE; {access Read Only}
   M211_M1_DR_IN_MAJ : MOTION_INSTRUCTION := (FLAGS := 570425344, DN := 1); {access None}
   M211_M1_DR_IN_MAM : MOTION_INSTRUCTION := (FLAGS := 33554432); {access None}
   M211_M1_DR_IN_MAR : MOTION_INSTRUCTION := (FLAGS := 33554432); {access None}
   M211_M1_DR_IN_MAS : MOTION_INSTRUCTION := (FLAGS := -1442840576, EN := 1, DN := 1, PC := 1); {access None}
   M211_M1_DR_IN_MCD : MOTION_INSTRUCTION := (FLAGS := 570425344, DN := 1); {access None}
   M211_M1_DR_IN_MRP : MOTION_INSTRUCTION := (FLAGS := 33554432); {access None}
   M211_M1_DR_MAFR : MOTION_INSTRUCTION := (FLAGS := 301989888, ER := 1, ERR := 11); {access None}
   M211_M1_DR_MDR : MOTION_INSTRUCTION := (FLAGS := -1845493760, EN := 1, ER := 1, ERR := 11); {access None}
   M211_M1_DR_MSF : MOTION_INSTRUCTION := (FLAGS := 570425344, DN := 1, STATUS := 2, STATE := 1); {access None}
   M211_M1_DR_MSO : MOTION_INSTRUCTION := (FLAGS := -1610612736, EN := 1, DN := 1, STATE := 1); {access None}
   M211_M1_DR_OUT_MAJ : MOTION_INSTRUCTION := (FLAGS := 570425344, DN := 1); {access None}
   M211_M1_DR_OUT_MAM : MOTION_INSTRUCTION := (FLAGS := 33554432); {access None}
   M211_M1_DR_OUT_MAR : MOTION_INSTRUCTION := (FLAGS := 33554432); {access None}
   M211_M1_DR_OUT_MAS : MOTION_INSTRUCTION := (FLAGS := -1442840576, EN := 1, DN := 1, PC := 1); {access None}
   M211_M1_DR_OUT_MCD : MOTION_INSTRUCTION := (FLAGS := 570425344, DN := 1); {access None}
   M211_M1_DR_OUT_MRP : MOTION_INSTRUCTION := (FLAGS := 33554432); {access None}
   M212_M1_DR : AXIS_CIP_DRIVE; {access Read Only}
   M212_M1_DR_IN_MAJ : MOTION_INSTRUCTION := (FLAGS := 570425344, DN := 1); {access None}
   M212_M1_DR_IN_MAM : MOTION_INSTRUCTION := (FLAGS := 33554432); {access None}
   M212_M1_DR_IN_MAR : MOTION_INSTRUCTION := (FLAGS := 33554432); {access None}
   M212_M1_DR_IN_MAS : MOTION_INSTRUCTION := (FLAGS := -1442840576, EN := 1, DN := 1, PC := 1); {access None}
   M212_M1_DR_IN_MCD : MOTION_INSTRUCTION := (FLAGS := 570425344, DN := 1); {access None}
   M212_M1_DR_IN_MRP : MOTION_INSTRUCTION := (FLAGS := 33554432); {access None}
   M212_M1_DR_MAFR : MOTION_INSTRUCTION := (FLAGS := 301989888, ER := 1, ERR := 11); {access None}
   M212_M1_DR_MDR : MOTION_INSTRUCTION := (FLAGS := -1845493760, EN := 1, ER := 1, ERR := 11); {access None}
